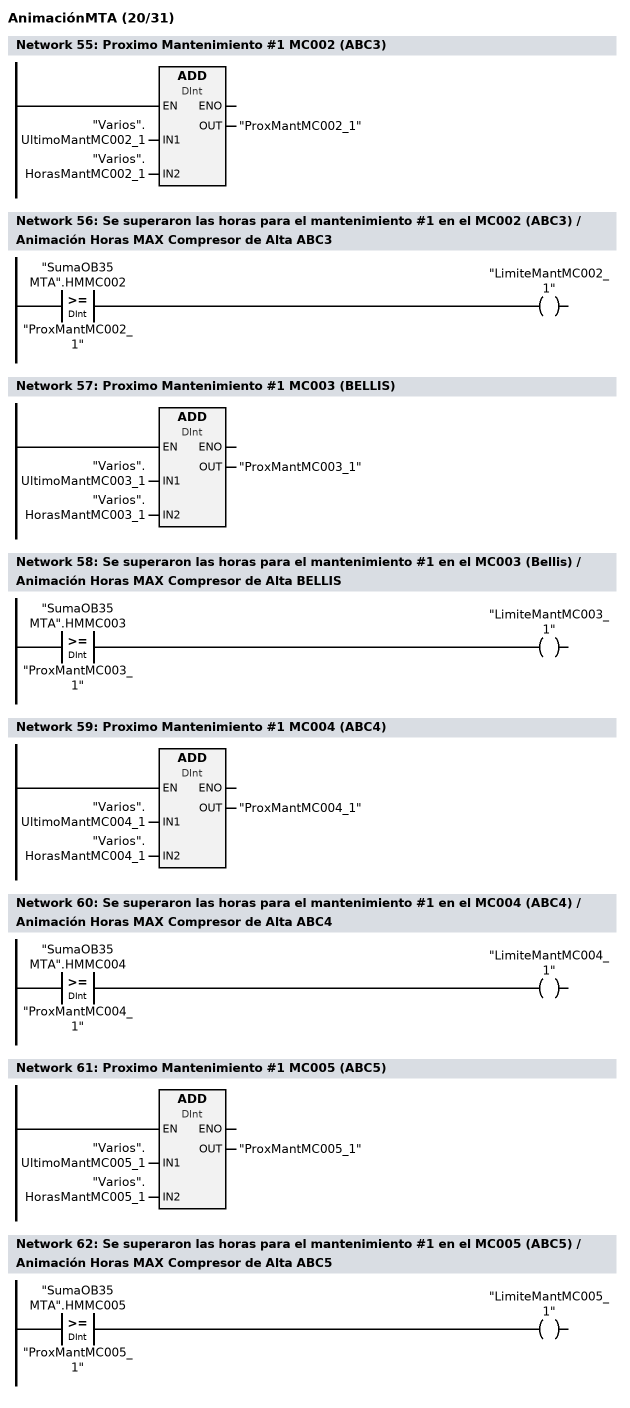
   RUNG wire#powerrail
      { S7_Templates := "SrcType := DInt"; S7_GenerateENO := "TRUE" } Add(in1 := "Varios".UltimoMantMC002_1, in2 := "Varios".HorasMantMC002_1, out => "ProxMantMC002_1")
   END_RUNG
   // the same network as SCL:
   "ProxMantMC002_1" := "Varios".UltimoMantMC002_1 + "Varios".HorasMantMC002_1;
END_REGION

REGION Network 56: Se superaron las horas para el mantenimiento #1 en el MC002 (ABC3) / Animación Horas MAX Compresor de Alta ABC3
   RUNG wire#powerrail
      { S7_Templates := "SrcType := DInt" } GE_Contact(in1 := "SumaOB35 MTA".HMMC002, in2 := "ProxMantMC002_1")
      Coil( "LimiteMantMC002_1" )
   END_RUNG
   // the same network as SCL:
   "LimiteMantMC002_1" := "SumaOB35 MTA".HMMC002 >= "ProxMantMC002_1";
END_REGION

REGION Network 57: Proximo Mantenimiento #1 MC003 (BELLIS)
   RUNG wire#powerrail
      { S7_Templates := "SrcType := DInt"; S7_GenerateENO := "TRUE" } Add(in1 := "Varios".UltimoMantMC003_1, in2 := "Varios".HorasMantMC003_1, out => "ProxMantMC003_1")
   END_RUNG
   // the same network as SCL:
   "ProxMantMC003_1" := "Varios".UltimoMantMC003_1 + "Varios".HorasMantMC003_1;
END_REGION

REGION Network 58: Se superaron las horas para el mantenimiento #1 en el MC003 (Bellis) / Animación Horas MAX Compresor de Alta BELLIS
   RUNG wire#powerrail
      { S7_Templates := "SrcType := DInt" } GE_Contact(in1 := "SumaOB35 MTA".HMMC003, in2 := "ProxMantMC003_1")
      Coil( "LimiteMantMC003_1" )
   END_RUNG
   // the same network as SCL:
   "LimiteMantMC003_1" := "SumaOB35 MTA".HMMC003 >= "ProxMantMC003_1";
END_REGION

REGION Network 59: Proximo Mantenimiento #1 MC004 (ABC4)
   RUNG wire#powerrail
      { S7_Templates := "SrcType := DInt"; S7_GenerateENO := "TRUE" } Add(in1 := "Varios".UltimoMantMC004_1, in2 := "Varios".HorasMantMC004_1, out => "ProxMantMC004_1")
   END_RUNG
   // the same network as SCL:
   "ProxMantMC004_1" := "Varios".UltimoMantMC004_1 + "Varios".HorasMantMC004_1;
END_REGION

REGION Network 60: Se superaron las horas para el mantenimiento #1 en el MC004 (ABC4) / Animación Horas MAX Compresor de Alta ABC4
   RUNG wire#powerrail
      { S7_Templates := "SrcType := DInt" } GE_Contact(in1 := "SumaOB35 MTA".HMMC004, in2 := "ProxMantMC004_1")
      Coil( "LimiteMantMC004_1" )
   END_RUNG
   // the same network as SCL:
   "LimiteMantMC004_1" := "SumaOB35 MTA".HMMC004 >= "ProxMantMC004_1";
END_REGION

REGION Network 61: Proximo Mantenimiento #1 MC005 (ABC5)
   RUNG wire#powerrail
      { S7_Templates := "SrcType := DInt"; S7_GenerateENO := "TRUE" } Add(in1 := "Varios".UltimoMantMC005_1, in2 := "Varios".HorasMantMC005_1, out => "ProxMantMC005_1")
   END_RUNG
   // the same network as SCL:
   "ProxMantMC005_1" := "Varios".UltimoMantMC005_1 + "Varios".HorasMantMC005_1;
END_REGION

REGION Network 62: Se superaron las horas para el mantenimiento #1 en el MC005 (ABC5) / Animación Horas MAX Compresor de Alta ABC5
   RUNG wire#powerrail
      { S7_Templates := "SrcType := DInt" } GE_Contact(in1 := "SumaOB35 MTA".HMMC005, in2 := "ProxMantMC005_1")
      Coil( "LimiteMantMC005_1" )
   END_RUNG
   // the same network as SCL:
   "LimiteMantMC005_1" := "SumaOB35 MTA".HMMC005 >= "ProxMantMC005_1";
END_REGION

REGION Network 63: Proximo Mantenimiento #1 MC006 (ABC1)
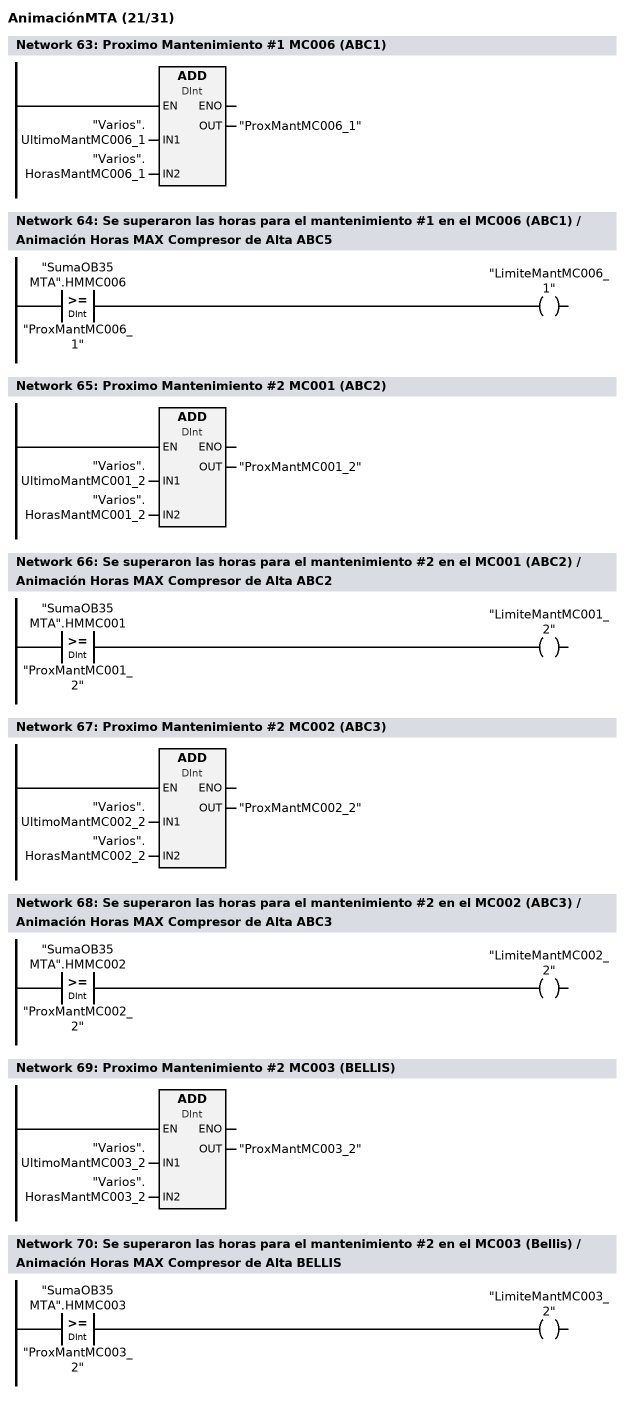
   RUNG wire#powerrail
      { S7_Templates := "SrcType := DInt"; S7_GenerateENO := "TRUE" } Add(in1 := "Varios".UltimoMantMC006_1, in2 := "Varios".HorasMantMC006_1, out => "ProxMantMC006_1")
   END_RUNG
   // the same network as SCL:
   "ProxMantMC006_1" := "Varios".UltimoMantMC006_1 + "Varios".HorasMantMC006_1;
END_REGION

REGION Network 64: Se superaron las horas para el mantenimiento #1 en el MC006 (ABC1) / Animación Horas MAX Compresor de Alta ABC5
   RUNG wire#powerrail
      { S7_Templates := "SrcType := DInt" } GE_Contact(in1 := "SumaOB35 MTA".HMMC006, in2 := "ProxMantMC006_1")
      Coil( "LimiteMantMC006_1" )
   END_RUNG
   // the same network as SCL:
   "LimiteMantMC006_1" := "SumaOB35 MTA".HMMC006 >= "ProxMantMC006_1";
END_REGION

REGION Network 65: Proximo Mantenimiento #2 MC001 (ABC2)
   RUNG wire#powerrail
      { S7_Templates := "SrcType := DInt"; S7_GenerateENO := "TRUE" } Add(in1 := "Varios".UltimoMantMC001_2, in2 := "Varios".HorasMantMC001_2, out => "ProxMantMC001_2")
   END_RUNG
   // the same network as SCL:
   "ProxMantMC001_2" := "Varios".UltimoMantMC001_2 + "Varios".HorasMantMC001_2;
END_REGION

REGION Network 66: Se superaron las horas para el mantenimiento #2 en el MC001 (ABC2) / Animación Horas MAX Compresor de Alta ABC2
   RUNG wire#powerrail
      { S7_Templates := "SrcType := DInt" } GE_Contact(in1 := "SumaOB35 MTA".HMMC001, in2 := "ProxMantMC001_2")
      Coil( "LimiteMantMC001_2" )
   END_RUNG
   // the same network as SCL:
   "LimiteMantMC001_2" := "SumaOB35 MTA".HMMC001 >= "ProxMantMC001_2";
END_REGION

REGION Network 67: Proximo Mantenimiento #2 MC002 (ABC3)
   RUNG wire#powerrail
      { S7_Templates := "SrcType := DInt"; S7_GenerateENO := "TRUE" } Add(in1 := "Varios".UltimoMantMC002_2, in2 := "Varios".HorasMantMC002_2, out => "ProxMantMC002_2")
   END_RUNG
   // the same network as SCL:
   "ProxMantMC002_2" := "Varios".UltimoMantMC002_2 + "Varios".HorasMantMC002_2;
END_REGION

REGION Network 68: Se superaron las horas para el mantenimiento #2 en el MC002 (ABC3) / Animación Horas MAX Compresor de Alta ABC3
   RUNG wire#powerrail
      { S7_Templates := "SrcType := DInt" } GE_Contact(in1 := "SumaOB35 MTA".HMMC002, in2 := "ProxMantMC002_2")
      Coil( "LimiteMantMC002_2" )
   END_RUNG
   // the same network as SCL:
   "LimiteMantMC002_2" := "SumaOB35 MTA".HMMC002 >= "ProxMantMC002_2";
END_REGION

REGION Network 69: Proximo Mantenimiento #2 MC003 (BELLIS)
   RUNG wire#powerrail
      { S7_Templates := "SrcType := DInt"; S7_GenerateENO := "TRUE" } Add(in1 := "Varios".UltimoMantMC003_2, in2 := "Varios".HorasMantMC003_2, out => "ProxMantMC003_2")
   END_RUNG
   // the same network as SCL:
   "ProxMantMC003_2" := "Varios".UltimoMantMC003_2 + "Varios".HorasMantMC003_2;
END_REGION

REGION Network 70: Se superaron las horas para el mantenimiento #2 en el MC003 (Bellis) / Animación Horas MAX Compresor de Alta BELLIS
   RUNG wire#powerrail
      { S7_Templates := "SrcType := DInt" } GE_Contact(in1 := "SumaOB35 MTA".HMMC003, in2 := "ProxMantMC003_2")
      Coil( "LimiteMantMC003_2" )
   END_RUNG
   // the same network as SCL:
   "LimiteMantMC003_2" := "SumaOB35 MTA".HMMC003 >= "ProxMantMC003_2";
END_REGION

REGION Network 71: Proximo Mantenimiento #2 MC004 (ABC4)
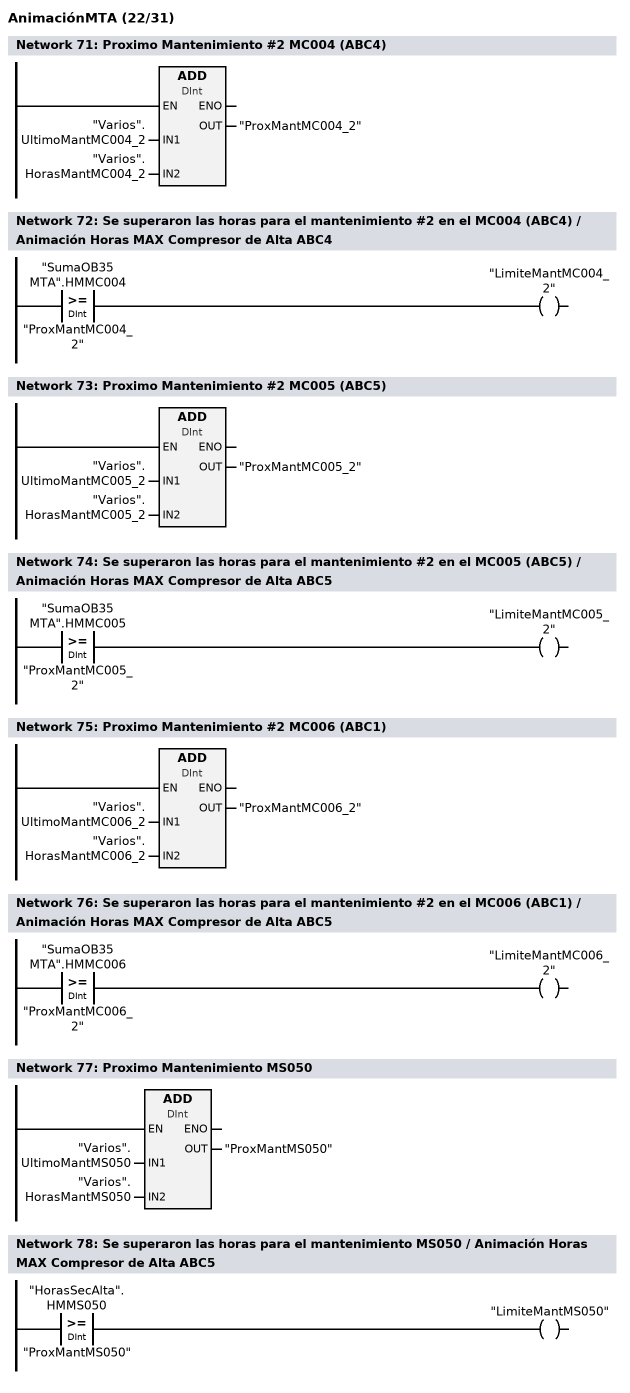
   RUNG wire#powerrail
      { S7_Templates := "SrcType := DInt"; S7_GenerateENO := "TRUE" } Add(in1 := "Varios".UltimoMantMC004_2, in2 := "Varios".HorasMantMC004_2, out => "ProxMantMC004_2")
   END_RUNG
   // the same network as SCL:
   "ProxMantMC004_2" := "Varios".UltimoMantMC004_2 + "Varios".HorasMantMC004_2;
END_REGION

REGION Network 72: Se superaron las horas para el mantenimiento #2 en el MC004 (ABC4) / Animación Horas MAX Compresor de Alta ABC4
   RUNG wire#powerrail
      { S7_Templates := "SrcType := DInt" } GE_Contact(in1 := "SumaOB35 MTA".HMMC004, in2 := "ProxMantMC004_2")
      Coil( "LimiteMantMC004_2" )
   END_RUNG
   // the same network as SCL:
   "LimiteMantMC004_2" := "SumaOB35 MTA".HMMC004 >= "ProxMantMC004_2";
END_REGION

REGION Network 73: Proximo Mantenimiento #2 MC005 (ABC5)
   RUNG wire#powerrail
      { S7_Templates := "SrcType := DInt"; S7_GenerateENO := "TRUE" } Add(in1 := "Varios".UltimoMantMC005_2, in2 := "Varios".HorasMantMC005_2, out => "ProxMantMC005_2")
   END_RUNG
   // the same network as SCL:
   "ProxMantMC005_2" := "Varios".UltimoMantMC005_2 + "Varios".HorasMantMC005_2;
END_REGION

REGION Network 74: Se superaron las horas para el mantenimiento #2 en el MC005 (ABC5) / Animación Horas MAX Compresor de Alta ABC5
   RUNG wire#powerrail
      { S7_Templates := "SrcType := DInt" } GE_Contact(in1 := "SumaOB35 MTA".HMMC005, in2 := "ProxMantMC005_2")
      Coil( "LimiteMantMC005_2" )
   END_RUNG
   // the same network as SCL:
   "LimiteMantMC005_2" := "SumaOB35 MTA".HMMC005 >= "ProxMantMC005_2";
END_REGION

REGION Network 75: Proximo Mantenimiento #2 MC006 (ABC1)
   RUNG wire#powerrail
      { S7_Templates := "SrcType := DInt"; S7_GenerateENO := "TRUE" } Add(in1 := "Varios".UltimoMantMC006_2, in2 := "Varios".HorasMantMC006_2, out => "ProxMantMC006_2")
   END_RUNG
   // the same network as SCL:
   "ProxMantMC006_2" := "Varios".UltimoMantMC006_2 + "Varios".HorasMantMC006_2;
END_REGION

REGION Network 76: Se superaron las horas para el mantenimiento #2 en el MC006 (ABC1) / Animación Horas MAX Compresor de Alta ABC5
   RUNG wire#powerrail
      { S7_Templates := "SrcType := DInt" } GE_Contact(in1 := "SumaOB35 MTA".HMMC006, in2 := "ProxMantMC006_2")
      Coil( "LimiteMantMC006_2" )
   END_RUNG
   // the same network as SCL:
   "LimiteMantMC006_2" := "SumaOB35 MTA".HMMC006 >= "ProxMantMC006_2";
END_REGION

REGION Network 77: Proximo Mantenimiento MS050
   RUNG wire#powerrail
      { S7_Templates := "SrcType := DInt"; S7_GenerateENO := "TRUE" } Add(in1 := "Varios".UltimoMantMS050, in2 := "Varios".HorasMantMS050, out => "ProxMantMS050")
   END_RUNG
   // the same network as SCL:
   "ProxMantMS050" := "Varios".UltimoMantMS050 + "Varios".HorasMantMS050;
END_REGION

REGION Network 78: Se superaron las horas para el mantenimiento MS050 / Animación Horas MAX Compresor de Alta ABC5
   RUNG wire#powerrail
      { S7_Templates := "SrcType := DInt" } GE_Contact(in1 := "HorasSecAlta".HMMS050, in2 := "ProxMantMS050")
      Coil( "LimiteMantMS050" )
   END_RUNG
   // the same network as SCL:
   "LimiteMantMS050" := "HorasSecAlta".HMMS050 >= "ProxMantMS050";
END_REGION

REGION Network 79: Proximo Mantenimiento MS051
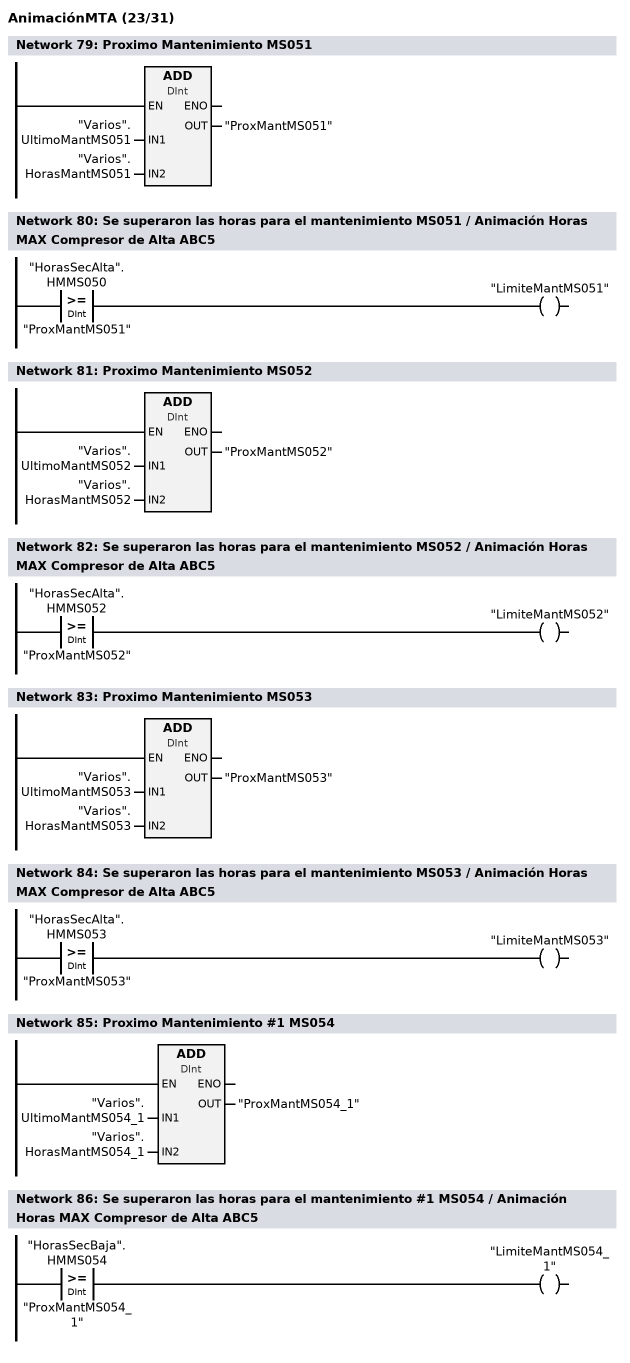
   RUNG wire#powerrail
      { S7_Templates := "SrcType := DInt"; S7_GenerateENO := "TRUE" } Add(in1 := "Varios".UltimoMantMS051, in2 := "Varios".HorasMantMS051, out => "ProxMantMS051")
   END_RUNG
   // the same network as SCL:
   "ProxMantMS051" := "Varios".UltimoMantMS051 + "Varios".HorasMantMS051;
END_REGION

REGION Network 80: Se superaron las horas para el mantenimiento MS051 / Animación Horas MAX Compresor de Alta ABC5
   RUNG wire#powerrail
      { S7_Templates := "SrcType := DInt" } GE_Contact(in1 := "HorasSecAlta".HMMS050, in2 := "ProxMantMS051")
      Coil( "LimiteMantMS051" )
   END_RUNG
   // the same network as SCL:
   "LimiteMantMS051" := "HorasSecAlta".HMMS050 >= "ProxMantMS051";
END_REGION

REGION Network 81: Proximo Mantenimiento MS052
   RUNG wire#powerrail
      { S7_Templates := "SrcType := DInt"; S7_GenerateENO := "TRUE" } Add(in1 := "Varios".UltimoMantMS052, in2 := "Varios".HorasMantMS052, out => "ProxMantMS052")
   END_RUNG
   // the same network as SCL:
   "ProxMantMS052" := "Varios".UltimoMantMS052 + "Varios".HorasMantMS052;
END_REGION

REGION Network 82: Se superaron las horas para el mantenimiento MS052 / Animación Horas MAX Compresor de Alta ABC5
   RUNG wire#powerrail
      { S7_Templates := "SrcType := DInt" } GE_Contact(in1 := "HorasSecAlta".HMMS052, in2 := "ProxMantMS052")
      Coil( "LimiteMantMS052" )
   END_RUNG
   // the same network as SCL:
   "LimiteMantMS052" := "HorasSecAlta".HMMS052 >= "ProxMantMS052";
END_REGION

REGION Network 83: Proximo Mantenimiento MS053
   RUNG wire#powerrail
      { S7_Templates := "SrcType := DInt"; S7_GenerateENO := "TRUE" } Add(in1 := "Varios".UltimoMantMS053, in2 := "Varios".HorasMantMS053, out => "ProxMantMS053")
   END_RUNG
   // the same network as SCL:
   "ProxMantMS053" := "Varios".UltimoMantMS053 + "Varios".HorasMantMS053;
END_REGION

REGION Network 84: Se superaron las horas para el mantenimiento MS053 / Animación Horas MAX Compresor de Alta ABC5
   RUNG wire#powerrail
      { S7_Templates := "SrcType := DInt" } GE_Contact(in1 := "HorasSecAlta".HMMS053, in2 := "ProxMantMS053")
      Coil( "LimiteMantMS053" )
   END_RUNG
   // the same network as SCL:
   "LimiteMantMS053" := "HorasSecAlta".HMMS053 >= "ProxMantMS053";
END_REGION

REGION Network 85: Proximo Mantenimiento #1 MS054
   RUNG wire#powerrail
      { S7_Templates := "SrcType := DInt"; S7_GenerateENO := "TRUE" } Add(in1 := "Varios".UltimoMantMS054_1, in2 := "Varios".HorasMantMS054_1, out => "ProxMantMS054_1")
   END_RUNG
   // the same network as SCL:
   "ProxMantMS054_1" := "Varios".UltimoMantMS054_1 + "Varios".HorasMantMS054_1;
END_REGION

REGION Network 86: Se superaron las horas para el mantenimiento #1 MS054 / Animación Horas MAX Compresor de Alta ABC5
   RUNG wire#powerrail
      { S7_Templates := "SrcType := DInt" } GE_Contact(in1 := "HorasSecBaja".HMMS054, in2 := "ProxMantMS054_1")
      Coil( "LimiteMantMS054_1" )
   END_RUNG
   // the same network as SCL:
   "LimiteMantMS054_1" := "HorasSecBaja".HMMS054 >= "ProxMantMS054_1";
END_REGION

REGION Network 87: Proximo Mantenimiento #2 MS054
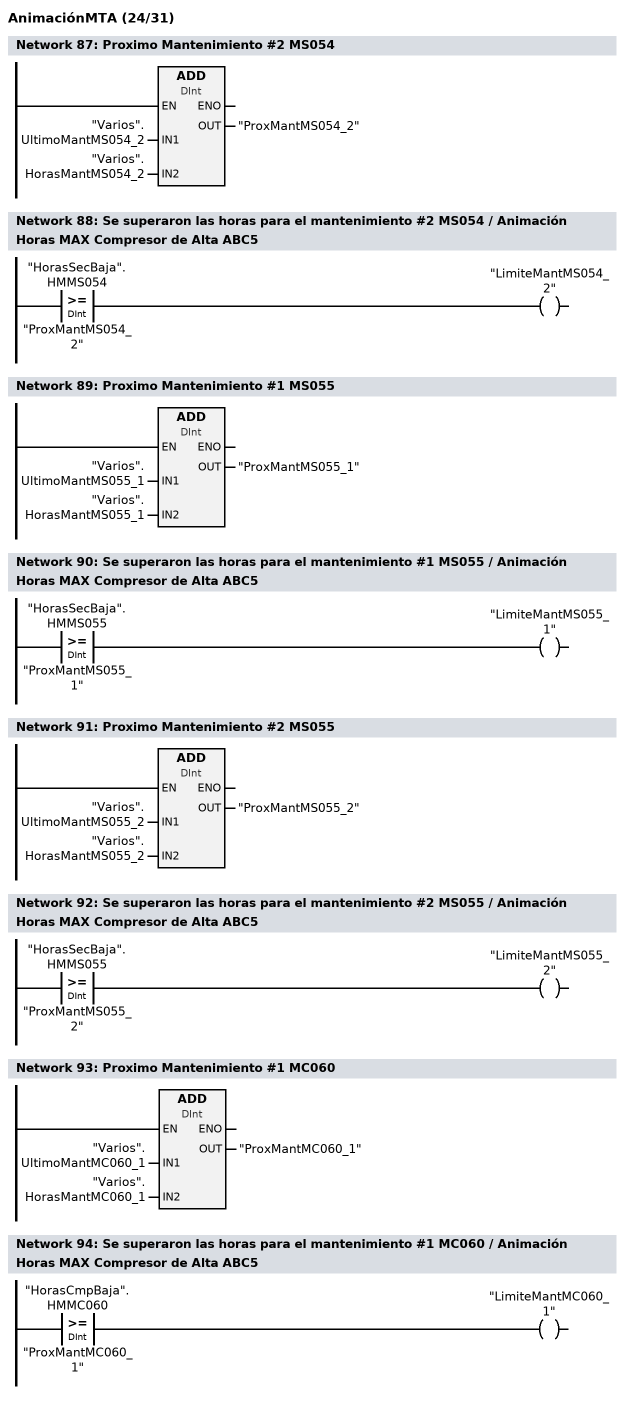
   RUNG wire#powerrail
      { S7_Templates := "SrcType := DInt"; S7_GenerateENO := "TRUE" } Add(in1 := "Varios".UltimoMantMS054_2, in2 := "Varios".HorasMantMS054_2, out => "ProxMantMS054_2")
   END_RUNG
   // the same network as SCL:
   "ProxMantMS054_2" := "Varios".UltimoMantMS054_2 + "Varios".HorasMantMS054_2;
END_REGION

REGION Network 88: Se superaron las horas para el mantenimiento #2 MS054 / Animación Horas MAX Compresor de Alta ABC5
   RUNG wire#powerrail
      { S7_Templates := "SrcType := DInt" } GE_Contact(in1 := "HorasSecBaja".HMMS054, in2 := "ProxMantMS054_2")
      Coil( "LimiteMantMS054_2" )
   END_RUNG
   // the same network as SCL:
   "LimiteMantMS054_2" := "HorasSecBaja".HMMS054 >= "ProxMantMS054_2";
END_REGION

REGION Network 89: Proximo Mantenimiento #1 MS055
   RUNG wire#powerrail
      { S7_Templates := "SrcType := DInt"; S7_GenerateENO := "TRUE" } Add(in1 := "Varios".UltimoMantMS055_1, in2 := "Varios".HorasMantMS055_1, out => "ProxMantMS055_1")
   END_RUNG
   // the same network as SCL:
   "ProxMantMS055_1" := "Varios".UltimoMantMS055_1 + "Varios".HorasMantMS055_1;
END_REGION

REGION Network 90: Se superaron las horas para el mantenimiento #1 MS055 / Animación Horas MAX Compresor de Alta ABC5
   RUNG wire#powerrail
      { S7_Templates := "SrcType := DInt" } GE_Contact(in1 := "HorasSecBaja".HMMS055, in2 := "ProxMantMS055_1")
      Coil( "LimiteMantMS055_1" )
   END_RUNG
   // the same network as SCL:
   "LimiteMantMS055_1" := "HorasSecBaja".HMMS055 >= "ProxMantMS055_1";
END_REGION

REGION Network 91: Proximo Mantenimiento #2 MS055
   RUNG wire#powerrail
      { S7_Templates := "SrcType := DInt"; S7_GenerateENO := "TRUE" } Add(in1 := "Varios".UltimoMantMS055_2, in2 := "Varios".HorasMantMS055_2, out => "ProxMantMS055_2")
   END_RUNG
   // the same network as SCL:
   "ProxMantMS055_2" := "Varios".UltimoMantMS055_2 + "Varios".HorasMantMS055_2;
END_REGION

REGION Network 92: Se superaron las horas para el mantenimiento #2 MS055 / Animación Horas MAX Compresor de Alta ABC5
   RUNG wire#powerrail
      { S7_Templates := "SrcType := DInt" } GE_Contact(in1 := "HorasSecBaja".HMMS055, in2 := "ProxMantMS055_2")
      Coil( "LimiteMantMS055_2" )
   END_RUNG
   // the same network as SCL:
   "LimiteMantMS055_2" := "HorasSecBaja".HMMS055 >= "ProxMantMS055_2";
END_REGION

REGION Network 93: Proximo Mantenimiento #1 MC060
   RUNG wire#powerrail
      { S7_Templates := "SrcType := DInt"; S7_GenerateENO := "TRUE" } Add(in1 := "Varios".UltimoMantMC060_1, in2 := "Varios".HorasMantMC060_1, out => "ProxMantMC060_1")
   END_RUNG
   // the same network as SCL:
   "ProxMantMC060_1" := "Varios".UltimoMantMC060_1 + "Varios".HorasMantMC060_1;
END_REGION

REGION Network 94: Se superaron las horas para el mantenimiento #1 MC060 / Animación Horas MAX Compresor de Alta ABC5
   RUNG wire#powerrail
      { S7_Templates := "SrcType := DInt" } GE_Contact(in1 := "HorasCmpBaja".HMMC060, in2 := "ProxMantMC060_1")
      Coil( "LimiteMantMC060_1" )
   END_RUNG
   // the same network as SCL:
   "LimiteMantMC060_1" := "HorasCmpBaja".HMMC060 >= "ProxMantMC060_1";
END_REGION

REGION Network 95: Proximo Mantenimiento #2 MC060
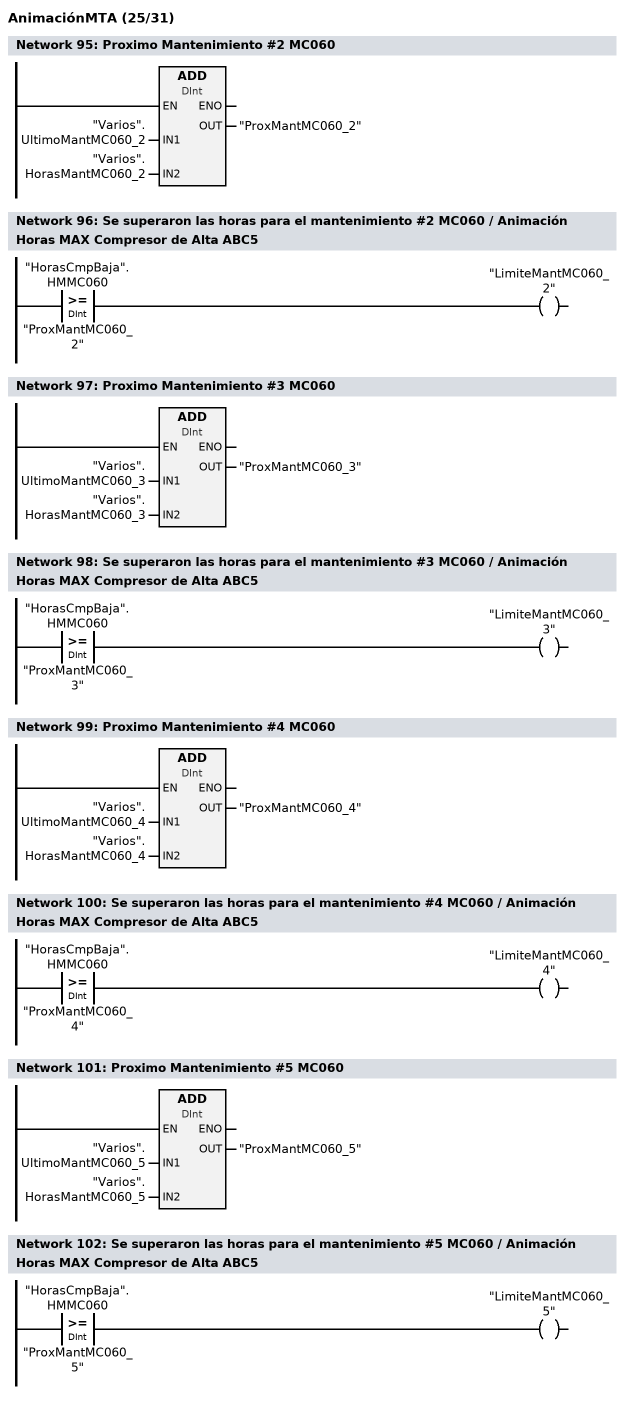
   RUNG wire#powerrail
      { S7_Templates := "SrcType := DInt"; S7_GenerateENO := "TRUE" } Add(in1 := "Varios".UltimoMantMC060_2, in2 := "Varios".HorasMantMC060_2, out => "ProxMantMC060_2")
   END_RUNG
   // the same network as SCL:
   "ProxMantMC060_2" := "Varios".UltimoMantMC060_2 + "Varios".HorasMantMC060_2;
END_REGION

REGION Network 96: Se superaron las horas para el mantenimiento #2 MC060 / Animación Horas MAX Compresor de Alta ABC5
   RUNG wire#powerrail
      { S7_Templates := "SrcType := DInt" } GE_Contact(in1 := "HorasCmpBaja".HMMC060, in2 := "ProxMantMC060_2")
      Coil( "LimiteMantMC060_2" )
   END_RUNG
   // the same network as SCL:
   "LimiteMantMC060_2" := "HorasCmpBaja".HMMC060 >= "ProxMantMC060_2";
END_REGION

REGION Network 97: Proximo Mantenimiento #3 MC060
   RUNG wire#powerrail
      { S7_Templates := "SrcType := DInt"; S7_GenerateENO := "TRUE" } Add(in1 := "Varios".UltimoMantMC060_3, in2 := "Varios".HorasMantMC060_3, out => "ProxMantMC060_3")
   END_RUNG
   // the same network as SCL:
   "ProxMantMC060_3" := "Varios".UltimoMantMC060_3 + "Varios".HorasMantMC060_3;
END_REGION

REGION Network 98: Se superaron las horas para el mantenimiento #3 MC060 / Animación Horas MAX Compresor de Alta ABC5
   RUNG wire#powerrail
      { S7_Templates := "SrcType := DInt" } GE_Contact(in1 := "HorasCmpBaja".HMMC060, in2 := "ProxMantMC060_3")
      Coil( "LimiteMantMC060_3" )
   END_RUNG
   // the same network as SCL:
   "LimiteMantMC060_3" := "HorasCmpBaja".HMMC060 >= "ProxMantMC060_3";
END_REGION

REGION Network 99: Proximo Mantenimiento #4 MC060
   RUNG wire#powerrail
      { S7_Templates := "SrcType := DInt"; S7_GenerateENO := "TRUE" } Add(in1 := "Varios".UltimoMantMC060_4, in2 := "Varios".HorasMantMC060_4, out => "ProxMantMC060_4")
   END_RUNG
   // the same network as SCL:
   "ProxMantMC060_4" := "Varios".UltimoMantMC060_4 + "Varios".HorasMantMC060_4;
END_REGION

REGION Network 100: Se superaron las horas para el mantenimiento #4 MC060 / Animación Horas MAX Compresor de Alta ABC5
   RUNG wire#powerrail
      { S7_Templates := "SrcType := DInt" } GE_Contact(in1 := "HorasCmpBaja".HMMC060, in2 := "ProxMantMC060_4")
      Coil( "LimiteMantMC060_4" )
   END_RUNG
   // the same network as SCL:
   "LimiteMantMC060_4" := "HorasCmpBaja".HMMC060 >= "ProxMantMC060_4";
END_REGION

REGION Network 101: Proximo Mantenimiento #5 MC060
   RUNG wire#powerrail
      { S7_Templates := "SrcType := DInt"; S7_GenerateENO := "TRUE" } Add(in1 := "Varios".UltimoMantMC060_5, in2 := "Varios".HorasMantMC060_5, out => "ProxMantMC060_5")
   END_RUNG
   // the same network as SCL:
   "ProxMantMC060_5" := "Varios".UltimoMantMC060_5 + "Varios".HorasMantMC060_5;
END_REGION

REGION Network 102: Se superaron las horas para el mantenimiento #5 MC060 / Animación Horas MAX Compresor de Alta ABC5
   RUNG wire#powerrail
      { S7_Templates := "SrcType := DInt" } GE_Contact(in1 := "HorasCmpBaja".HMMC060, in2 := "ProxMantMC060_5")
      Coil( "LimiteMantMC060_5" )
   END_RUNG
   // the same network as SCL:
   "LimiteMantMC060_5" := "HorasCmpBaja".HMMC060 >= "ProxMantMC060_5";
END_REGION

REGION Network 103: Proximo Mantenimiento #1 MC061
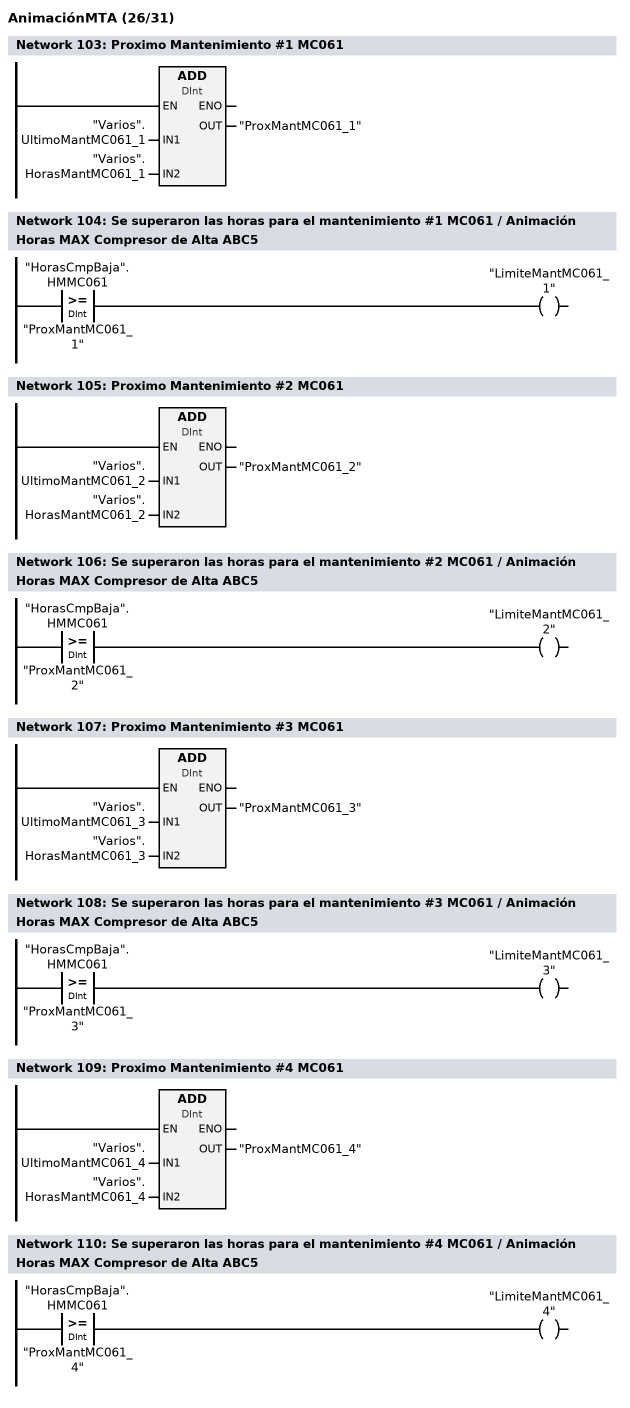
   RUNG wire#powerrail
      { S7_Templates := "SrcType := DInt"; S7_GenerateENO := "TRUE" } Add(in1 := "Varios".UltimoMantMC061_1, in2 := "Varios".HorasMantMC061_1, out => "ProxMantMC061_1")
   END_RUNG
   // the same network as SCL:
   "ProxMantMC061_1" := "Varios".UltimoMantMC061_1 + "Varios".HorasMantMC061_1;
END_REGION

REGION Network 104: Se superaron las horas para el mantenimiento #1 MC061 / Animación Horas MAX Compresor de Alta ABC5
   RUNG wire#powerrail
      { S7_Templates := "SrcType := DInt" } GE_Contact(in1 := "HorasCmpBaja".HMMC061, in2 := "ProxMantMC061_1")
      Coil( "LimiteMantMC061_1" )
   END_RUNG
   // the same network as SCL:
   "LimiteMantMC061_1" := "HorasCmpBaja".HMMC061 >= "ProxMantMC061_1";
END_REGION

REGION Network 105: Proximo Mantenimiento #2 MC061
   RUNG wire#powerrail
      { S7_Templates := "SrcType := DInt"; S7_GenerateENO := "TRUE" } Add(in1 := "Varios".UltimoMantMC061_2, in2 := "Varios".HorasMantMC061_2, out => "ProxMantMC061_2")
   END_RUNG
   // the same network as SCL:
   "ProxMantMC061_2" := "Varios".UltimoMantMC061_2 + "Varios".HorasMantMC061_2;
END_REGION

REGION Network 106: Se superaron las horas para el mantenimiento #2 MC061 / Animación Horas MAX Compresor de Alta ABC5
   RUNG wire#powerrail
      { S7_Templates := "SrcType := DInt" } GE_Contact(in1 := "HorasCmpBaja".HMMC061, in2 := "ProxMantMC061_2")
      Coil( "LimiteMantMC061_2" )
   END_RUNG
   // the same network as SCL:
   "LimiteMantMC061_2" := "HorasCmpBaja".HMMC061 >= "ProxMantMC061_2";
END_REGION

REGION Network 107: Proximo Mantenimiento #3 MC061
   RUNG wire#powerrail
      { S7_Templates := "SrcType := DInt"; S7_GenerateENO := "TRUE" } Add(in1 := "Varios".UltimoMantMC061_3, in2 := "Varios".HorasMantMC061_3, out => "ProxMantMC061_3")
   END_RUNG
   // the same network as SCL:
   "ProxMantMC061_3" := "Varios".UltimoMantMC061_3 + "Varios".HorasMantMC061_3;
END_REGION

REGION Network 108: Se superaron las horas para el mantenimiento #3 MC061 / Animación Horas MAX Compresor de Alta ABC5
   RUNG wire#powerrail
      { S7_Templates := "SrcType := DInt" } GE_Contact(in1 := "HorasCmpBaja".HMMC061, in2 := "ProxMantMC061_3")
      Coil( "LimiteMantMC061_3" )
   END_RUNG
   // the same network as SCL:
   "LimiteMantMC061_3" := "HorasCmpBaja".HMMC061 >= "ProxMantMC061_3";
END_REGION

REGION Network 109: Proximo Mantenimiento #4 MC061
   RUNG wire#powerrail
      { S7_Templates := "SrcType := DInt"; S7_GenerateENO := "TRUE" } Add(in1 := "Varios".UltimoMantMC061_4, in2 := "Varios".HorasMantMC061_4, out => "ProxMantMC061_4")
   END_RUNG
   // the same network as SCL:
   "ProxMantMC061_4" := "Varios".UltimoMantMC061_4 + "Varios".HorasMantMC061_4;
END_REGION

REGION Network 110: Se superaron las horas para el mantenimiento #4 MC061 / Animación Horas MAX Compresor de Alta ABC5
   RUNG wire#powerrail
      { S7_Templates := "SrcType := DInt" } GE_Contact(in1 := "HorasCmpBaja".HMMC061, in2 := "ProxMantMC061_4")
      Coil( "LimiteMantMC061_4" )
   END_RUNG
   // the same network as SCL:
   "LimiteMantMC061_4" := "HorasCmpBaja".HMMC061 >= "ProxMantMC061_4";
END_REGION

REGION Network 111: Proximo Mantenimiento #5 MC061
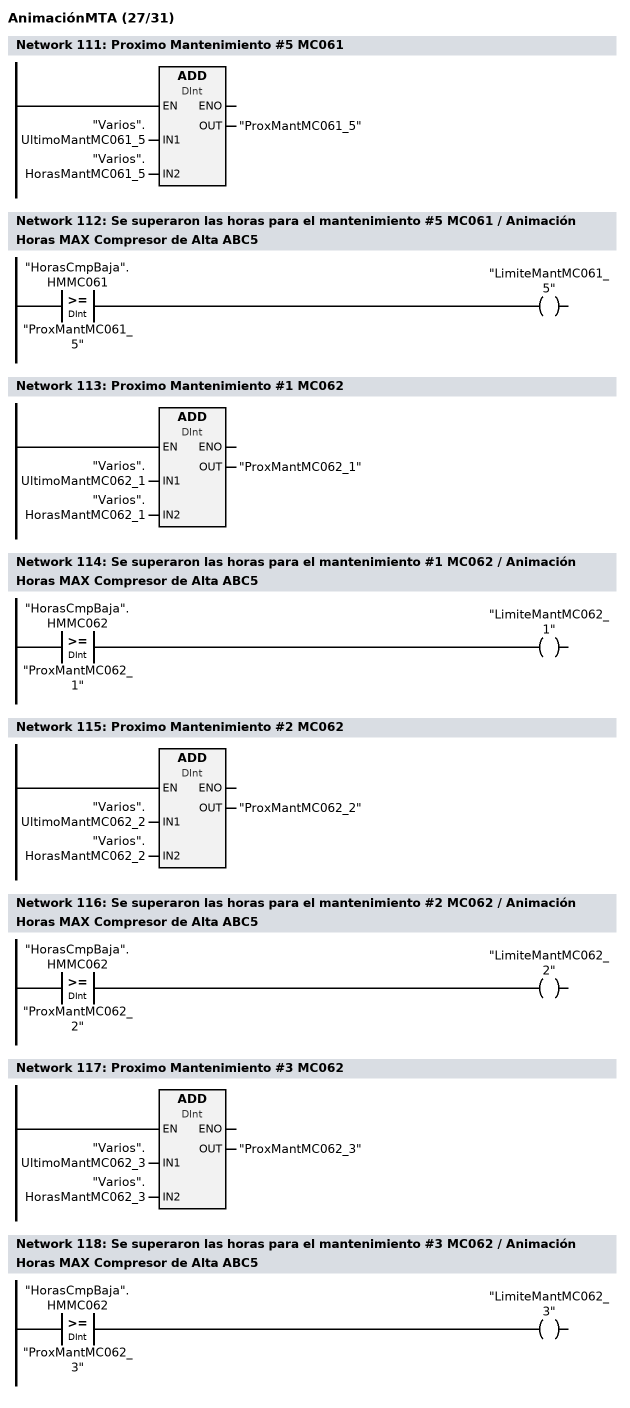
   RUNG wire#powerrail
      { S7_Templates := "SrcType := DInt"; S7_GenerateENO := "TRUE" } Add(in1 := "Varios".UltimoMantMC061_5, in2 := "Varios".HorasMantMC061_5, out => "ProxMantMC061_5")
   END_RUNG
   // the same network as SCL:
   "ProxMantMC061_5" := "Varios".UltimoMantMC061_5 + "Varios".HorasMantMC061_5;
END_REGION

REGION Network 112: Se superaron las horas para el mantenimiento #5 MC061 / Animación Horas MAX Compresor de Alta ABC5
   RUNG wire#powerrail
      { S7_Templates := "SrcType := DInt" } GE_Contact(in1 := "HorasCmpBaja".HMMC061, in2 := "ProxMantMC061_5")
      Coil( "LimiteMantMC061_5" )
   END_RUNG
   // the same network as SCL:
   "LimiteMantMC061_5" := "HorasCmpBaja".HMMC061 >= "ProxMantMC061_5";
END_REGION

REGION Network 113: Proximo Mantenimiento #1 MC062
   RUNG wire#powerrail
      { S7_Templates := "SrcType := DInt"; S7_GenerateENO := "TRUE" } Add(in1 := "Varios".UltimoMantMC062_1, in2 := "Varios".HorasMantMC062_1, out => "ProxMantMC062_1")
   END_RUNG
   // the same network as SCL:
   "ProxMantMC062_1" := "Varios".UltimoMantMC062_1 + "Varios".HorasMantMC062_1;
END_REGION

REGION Network 114: Se superaron las horas para el mantenimiento #1 MC062 / Animación Horas MAX Compresor de Alta ABC5
   RUNG wire#powerrail
      { S7_Templates := "SrcType := DInt" } GE_Contact(in1 := "HorasCmpBaja".HMMC062, in2 := "ProxMantMC062_1")
      Coil( "LimiteMantMC062_1" )
   END_RUNG
   // the same network as SCL:
   "LimiteMantMC062_1" := "HorasCmpBaja".HMMC062 >= "ProxMantMC062_1";
END_REGION

REGION Network 115: Proximo Mantenimiento #2 MC062
   RUNG wire#powerrail
      { S7_Templates := "SrcType := DInt"; S7_GenerateENO := "TRUE" } Add(in1 := "Varios".UltimoMantMC062_2, in2 := "Varios".HorasMantMC062_2, out => "ProxMantMC062_2")
   END_RUNG
   // the same network as SCL:
   "ProxMantMC062_2" := "Varios".UltimoMantMC062_2 + "Varios".HorasMantMC062_2;
END_REGION

REGION Network 116: Se superaron las horas para el mantenimiento #2 MC062 / Animación Horas MAX Compresor de Alta ABC5
   RUNG wire#powerrail
      { S7_Templates := "SrcType := DInt" } GE_Contact(in1 := "HorasCmpBaja".HMMC062, in2 := "ProxMantMC062_2")
      Coil( "LimiteMantMC062_2" )
   END_RUNG
   // the same network as SCL:
   "LimiteMantMC062_2" := "HorasCmpBaja".HMMC062 >= "ProxMantMC062_2";
END_REGION

REGION Network 117: Proximo Mantenimiento #3 MC062
   RUNG wire#powerrail
      { S7_Templates := "SrcType := DInt"; S7_GenerateENO := "TRUE" } Add(in1 := "Varios".UltimoMantMC062_3, in2 := "Varios".HorasMantMC062_3, out => "ProxMantMC062_3")
   END_RUNG
   // the same network as SCL:
   "ProxMantMC062_3" := "Varios".UltimoMantMC062_3 + "Varios".HorasMantMC062_3;
END_REGION

REGION Network 118: Se superaron las horas para el mantenimiento #3 MC062 / Animación Horas MAX Compresor de Alta ABC5
   RUNG wire#powerrail
      { S7_Templates := "SrcType := DInt" } GE_Contact(in1 := "HorasCmpBaja".HMMC062, in2 := "ProxMantMC062_3")
      Coil( "LimiteMantMC062_3" )
   END_RUNG
   // the same network as SCL:
   "LimiteMantMC062_3" := "HorasCmpBaja".HMMC062 >= "ProxMantMC062_3";
END_REGION

REGION Network 119: Proximo Mantenimiento #4 MC062